REGION Network 83
   RUNG wire#powerrail
      Move(in := "Carrier_54_G120DControlWord", out1 => "DB402_SDC_CARRIER_DRIVE_DATA".Drive_Data.CARRIER[54].Drive_Control)
      Move(in := "Carrier_54_G120DStatusWord", out1 => "DB402_SDC_CARRIER_DRIVE_DATA".Drive_Data.CARRIER[54].Drive_Status)
   END_RUNG
   // the same network as SCL:
   "DB402_SDC_CARRIER_DRIVE_DATA".Drive_Data.CARRIER[54].Drive_Control := "Carrier_54_G120DControlWord";
   "DB402_SDC_CARRIER_DRIVE_DATA".Drive_Data.CARRIER[54].Drive_Status := "Carrier_54_G120DStatusWord";
END_REGION

REGION Network 84
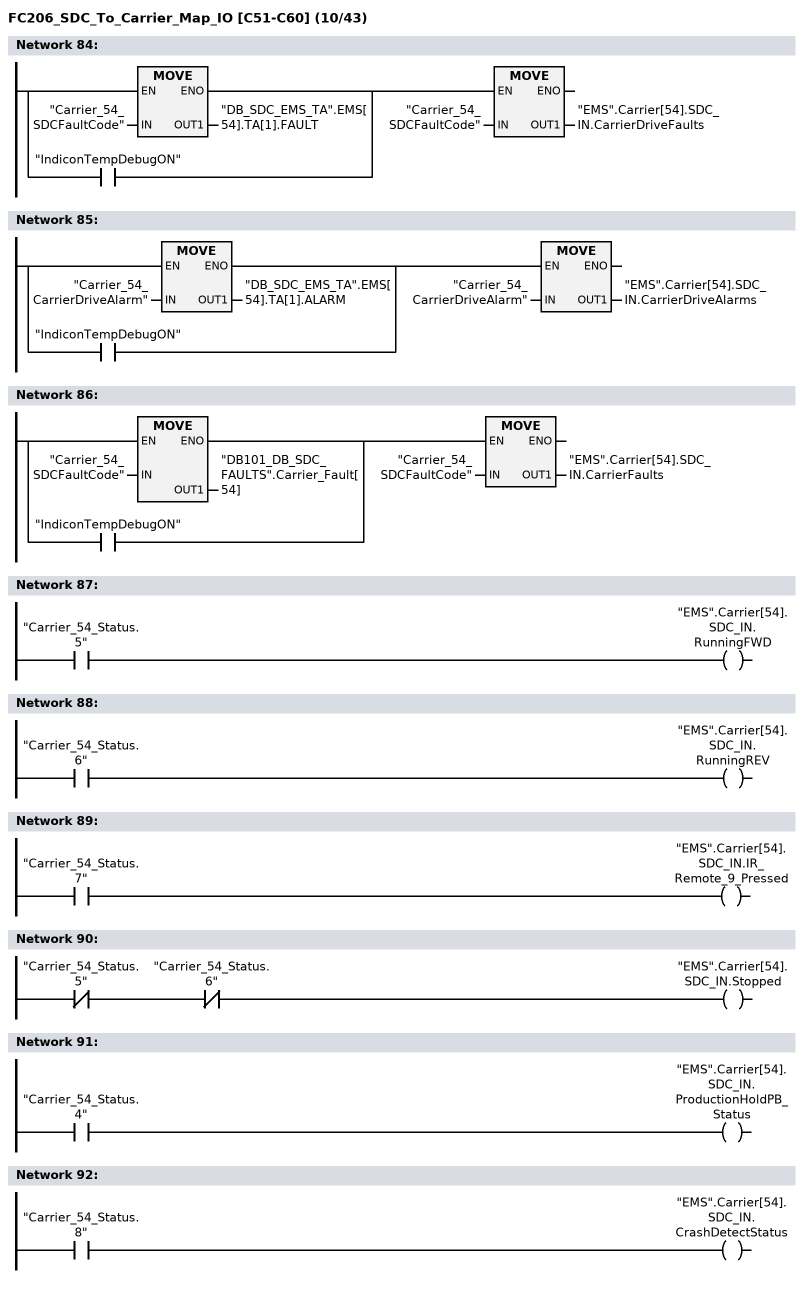
   RUNG wire#powerrail
      Move(in := "Carrier_54_SDCFaultCode", out1 => "DB_SDC_EMS_TA".EMS[54].TA[1].FAULT)
      wire#w1
      Move(in := "Carrier_54_SDCFaultCode", out1 => "EMS".Carrier[54].SDC_IN.CarrierDriveFaults)
   END_RUNG
   RUNG wire#powerrail
      Contact( "IndiconTempDebugON" )
   END_RUNG wire#w1
   // the same network as SCL:
   "DB_SDC_EMS_TA".EMS[54].TA[1].FAULT := "Carrier_54_SDCFaultCode";
   IF TRUE OR "IndiconTempDebugON" THEN
       "EMS".Carrier[54].SDC_IN.CarrierDriveFaults := "Carrier_54_SDCFaultCode";
   END_IF;
END_REGION

REGION Network 85
   RUNG wire#powerrail
      Move(in := "Carrier_54_CarrierDriveAlarm", out1 => "DB_SDC_EMS_TA".EMS[54].TA[1].ALARM)
      wire#w1
      Move(in := "Carrier_54_CarrierDriveAlarm", out1 => "EMS".Carrier[54].SDC_IN.CarrierDriveAlarms)
   END_RUNG
   RUNG wire#powerrail
      Contact( "IndiconTempDebugON" )
   END_RUNG wire#w1
   // the same network as SCL:
   "DB_SDC_EMS_TA".EMS[54].TA[1].ALARM := "Carrier_54_CarrierDriveAlarm";
   IF TRUE OR "IndiconTempDebugON" THEN
       "EMS".Carrier[54].SDC_IN.CarrierDriveAlarms := "Carrier_54_CarrierDriveAlarm";
   END_IF;
END_REGION

REGION Network 86
   RUNG wire#powerrail
      Move(in := "Carrier_54_SDCFaultCode", out1 => "DB101_DB_SDC_FAULTS".Carrier_Fault[54])
      wire#w1
      Move(in := "Carrier_54_SDCFaultCode", out1 => "EMS".Carrier[54].SDC_IN.CarrierFaults)
   END_RUNG
   RUNG wire#powerrail
      Contact( "IndiconTempDebugON" )
   END_RUNG wire#w1
   // the same network as SCL:
   "DB101_DB_SDC_FAULTS".Carrier_Fault[54] := "Carrier_54_SDCFaultCode";
   IF TRUE OR "IndiconTempDebugON" THEN
       "EMS".Carrier[54].SDC_IN.CarrierFaults := "Carrier_54_SDCFaultCode";
   END_IF;
END_REGION

REGION Network 87
   RUNG wire#powerrail
      Contact( "Carrier_54_Status.5" )
      Coil( "EMS".Carrier[54].SDC_IN.RunningFWD )
   END_RUNG
   // the same network as SCL:
   "EMS".Carrier[54].SDC_IN.RunningFWD := "Carrier_54_Status.5";
END_REGION

REGION Network 88
   RUNG wire#powerrail
      Contact( "Carrier_54_Status.6" )
      Coil( "EMS".Carrier[54].SDC_IN.RunningREV )
   END_RUNG
   // the same network as SCL:
   "EMS".Carrier[54].SDC_IN.RunningREV := "Carrier_54_Status.6";
END_REGION

REGION Network 89
   RUNG wire#powerrail
      Contact( "Carrier_54_Status.7" )
      Coil( "EMS".Carrier[54].SDC_IN.IR_Remote_9_Pressed )
   END_RUNG
   // the same network as SCL:
   "EMS".Carrier[54].SDC_IN.IR_Remote_9_Pressed := "Carrier_54_Status.7";
END_REGION

REGION Network 90
   RUNG wire#powerrail
      I_Contact( "Carrier_54_Status.5" )
      I_Contact( "Carrier_54_Status.6" )
      Coil( "EMS".Carrier[54].SDC_IN.Stopped )
   END_RUNG
   // the same network as SCL:
   "EMS".Carrier[54].SDC_IN.Stopped := NOT "Carrier_54_Status.5" AND NOT "Carrier_54_Status.6";
END_REGION

REGION Network 91
   RUNG wire#powerrail
      Contact( "Carrier_54_Status.4" )
      Coil( "EMS".Carrier[54].SDC_IN.ProductionHoldPB_Status )
   END_RUNG
   // the same network as SCL:
   "EMS".Carrier[54].SDC_IN.ProductionHoldPB_Status := "Carrier_54_Status.4";
END_REGION

REGION Network 92
   RUNG wire#powerrail
      Contact( "Carrier_54_Status.8" )
      Coil( "EMS".Carrier[54].SDC_IN.CrashDetectStatus )
   END_RUNG
   // the same network as SCL:
   "EMS".Carrier[54].SDC_IN.CrashDetectStatus := "Carrier_54_Status.8";
END_REGION

REGION Network 93
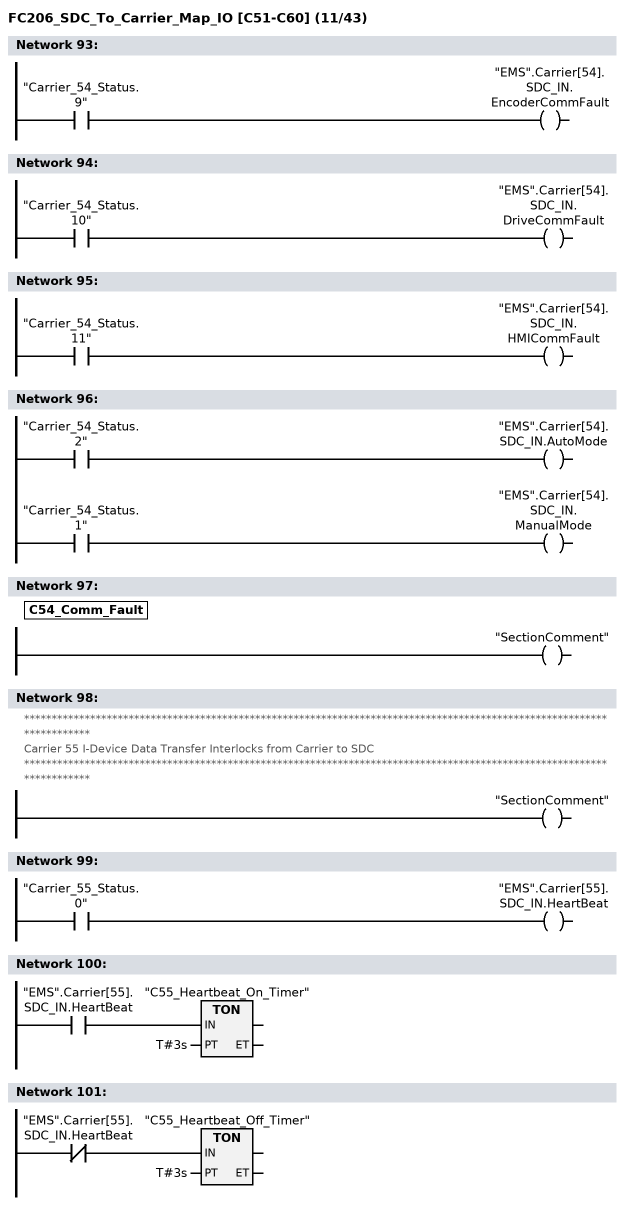
   RUNG wire#powerrail
      Contact( "Carrier_54_Status.9" )
      Coil( "EMS".Carrier[54].SDC_IN.EncoderCommFault )
   END_RUNG
   // the same network as SCL:
   "EMS".Carrier[54].SDC_IN.EncoderCommFault := "Carrier_54_Status.9";
END_REGION

REGION Network 94
   RUNG wire#powerrail
      Contact( "Carrier_54_Status.10" )
      Coil( "EMS".Carrier[54].SDC_IN.DriveCommFault )
   END_RUNG
   // the same network as SCL:
   "EMS".Carrier[54].SDC_IN.DriveCommFault := "Carrier_54_Status.10";
END_REGION

REGION Network 95
   RUNG wire#powerrail
      Contact( "Carrier_54_Status.11" )
      Coil( "EMS".Carrier[54].SDC_IN.HMICommFault )
   END_RUNG
   // the same network as SCL:
   "EMS".Carrier[54].SDC_IN.HMICommFault := "Carrier_54_Status.11";
END_REGION

REGION Network 96
   RUNG wire#powerrail
      Contact( "Carrier_54_Status.2" )
      Coil( "EMS".Carrier[54].SDC_IN.AutoMode )
   END_RUNG
   RUNG wire#powerrail
      Contact( "Carrier_54_Status.1" )
      Coil( "EMS".Carrier[54].SDC_IN.ManualMode )
   END_RUNG
   // the same network as SCL:
   "EMS".Carrier[54].SDC_IN.AutoMode := "Carrier_54_Status.2";
   "EMS".Carrier[54].SDC_IN.ManualMode := "Carrier_54_Status.1";
END_REGION

REGION Network 97
   Label( C54_Comm_Fault )
   RUNG wire#powerrail
      Coil( "SectionComment" )
   END_RUNG
   // the same network as SCL:
   C54_Comm_Fault:
   "SectionComment" := TRUE;
END_REGION

REGION Network 98
   // **********************************************************************************************************************
   // 
   // Carrier 55 I-Device Data Transfer Interlocks from Carrier to SDC
   // 
   // **********************************************************************************************************************
   RUNG wire#powerrail
      Coil( "SectionComment" )
   END_RUNG
   // the same network as SCL:
   "SectionComment" := TRUE;
END_REGION

REGION Network 99
   RUNG wire#powerrail
      Contact( "Carrier_55_Status.0" )
      Coil( "EMS".Carrier[55].SDC_IN.HeartBeat )
   END_RUNG
   // the same network as SCL:
   "EMS".Carrier[55].SDC_IN.HeartBeat := "Carrier_55_Status.0";
END_REGION

REGION Network 100
   "C55_Heartbeat_On_Timer".TON(IN := "EMS".Carrier[55].SDC_IN.HeartBeat, PT := T#3s);
END_REGION

REGION Network 101
   "C55_Heartbeat_Off_Timer".TON(IN := NOT "EMS".Carrier[55].SDC_IN.HeartBeat, PT := T#3s);
END_REGION

REGION Network 102
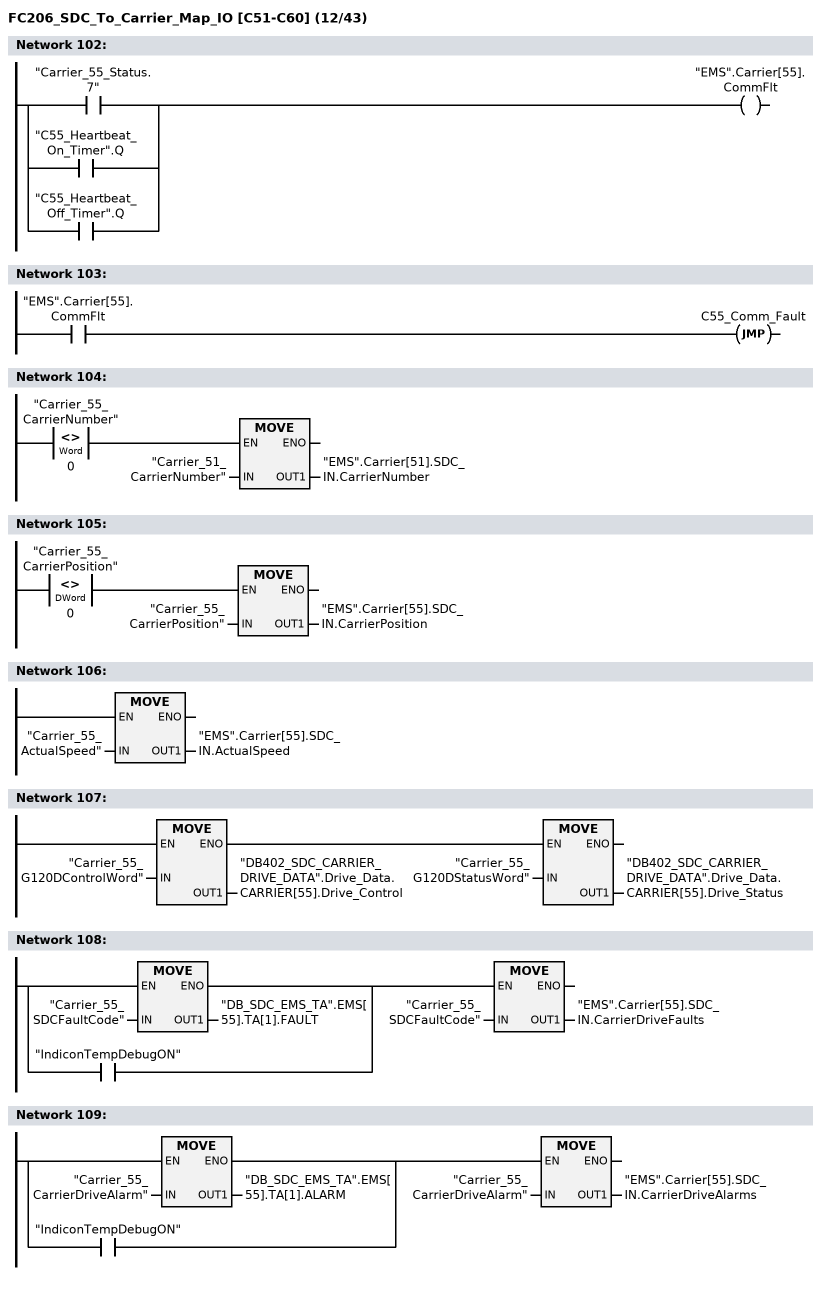
   RUNG wire#powerrail
      Contact( "Carrier_55_Status.7" )
      wire#w1
      Coil( "EMS".Carrier[55].CommFlt )
   END_RUNG
   RUNG wire#powerrail
      Contact( "C55_Heartbeat_On_Timer".Q )
   END_RUNG wire#w1
   RUNG wire#powerrail
      Contact( "C55_Heartbeat_Off_Timer".Q )
   END_RUNG wire#w1
   // the same network as SCL:
   "EMS".Carrier[55].CommFlt := "Carrier_55_Status.7" OR "C55_Heartbeat_On_Timer".Q OR "C55_Heartbeat_Off_Timer".Q;
END_REGION

REGION Network 103
   RUNG wire#powerrail
      Contact( "EMS".Carrier[55].CommFlt )
      JumpCoil( C55_Comm_Fault )
   END_RUNG
   // the same network as SCL:
   IF "EMS".Carrier[55].CommFlt THEN GOTO C55_Comm_Fault; END_IF;
END_REGION

REGION Network 104
   RUNG wire#powerrail
      { S7_Templates := "SrcType := Word" } NE_Contact(in1 := "Carrier_55_CarrierNumber", in2 := 0)
      Move(in := "Carrier_51_CarrierNumber", out1 => "EMS".Carrier[51].SDC_IN.CarrierNumber)
   END_RUNG
   // the same network as SCL:
   IF "Carrier_55_CarrierNumber" <> 0 THEN
       "EMS".Carrier[51].SDC_IN.CarrierNumber := "Carrier_51_CarrierNumber";
   END_IF;
END_REGION

REGION Network 105
   RUNG wire#powerrail
      { S7_Templates := "SrcType := DWord" } NE_Contact(in1 := "Carrier_55_CarrierPosition", in2 := 0)
      Move(in := "Carrier_55_CarrierPosition", out1 => "EMS".Carrier[55].SDC_IN.CarrierPosition)
   END_RUNG
   // the same network as SCL:
   IF "Carrier_55_CarrierPosition" <> 0 THEN
       "EMS".Carrier[55].SDC_IN.CarrierPosition := "Carrier_55_CarrierPosition";
   END_IF;
END_REGION

REGION Network 106
   RUNG wire#powerrail
      Move(in := "Carrier_55_ActualSpeed", out1 => "EMS".Carrier[55].SDC_IN.ActualSpeed)
   END_RUNG
   // the same network as SCL:
   "EMS".Carrier[55].SDC_IN.ActualSpeed := "Carrier_55_ActualSpeed";
END_REGION

REGION Network 107
   RUNG wire#powerrail
      Move(in := "Carrier_55_G120DControlWord", out1 => "DB402_SDC_CARRIER_DRIVE_DATA".Drive_Data.CARRIER[55].Drive_Control)
      Move(in := "Carrier_55_G120DStatusWord", out1 => "DB402_SDC_CARRIER_DRIVE_DATA".Drive_Data.CARRIER[55].Drive_Status)
   END_RUNG
   // the same network as SCL:
   "DB402_SDC_CARRIER_DRIVE_DATA".Drive_Data.CARRIER[55].Drive_Control := "Carrier_55_G120DControlWord";
   "DB402_SDC_CARRIER_DRIVE_DATA".Drive_Data.CARRIER[55].Drive_Status := "Carrier_55_G120DStatusWord";
END_REGION

REGION Network 108
   RUNG wire#powerrail
      Move(in := "Carrier_55_SDCFaultCode", out1 => "DB_SDC_EMS_TA".EMS[55].TA[1].FAULT)
      wire#w1
      Move(in := "Carrier_55_SDCFaultCode", out1 => "EMS".Carrier[55].SDC_IN.CarrierDriveFaults)
   END_RUNG
   RUNG wire#powerrail
      Contact( "IndiconTempDebugON" )
   END_RUNG wire#w1
   // the same network as SCL:
   "DB_SDC_EMS_TA".EMS[55].TA[1].FAULT := "Carrier_55_SDCFaultCode";
   IF TRUE OR "IndiconTempDebugON" THEN
       "EMS".Carrier[55].SDC_IN.CarrierDriveFaults := "Carrier_55_SDCFaultCode";
   END_IF;
END_REGION

REGION Network 109
   RUNG wire#powerrail
      Move(in := "Carrier_55_CarrierDriveAlarm", out1 => "DB_SDC_EMS_TA".EMS[55].TA[1].ALARM)
      wire#w1
      Move(in := "Carrier_55_CarrierDriveAlarm", out1 => "EMS".Carrier[55].SDC_IN.CarrierDriveAlarms)
   END_RUNG
   RUNG wire#powerrail
      Contact( "IndiconTempDebugON" )
   END_RUNG wire#w1
   // the same network as SCL:
   "DB_SDC_EMS_TA".EMS[55].TA[1].ALARM := "Carrier_55_CarrierDriveAlarm";
   IF TRUE OR "IndiconTempDebugON" THEN
       "EMS".Carrier[55].SDC_IN.CarrierDriveAlarms := "Carrier_55_CarrierDriveAlarm";
   END_IF;
END_REGION

REGION Network 110
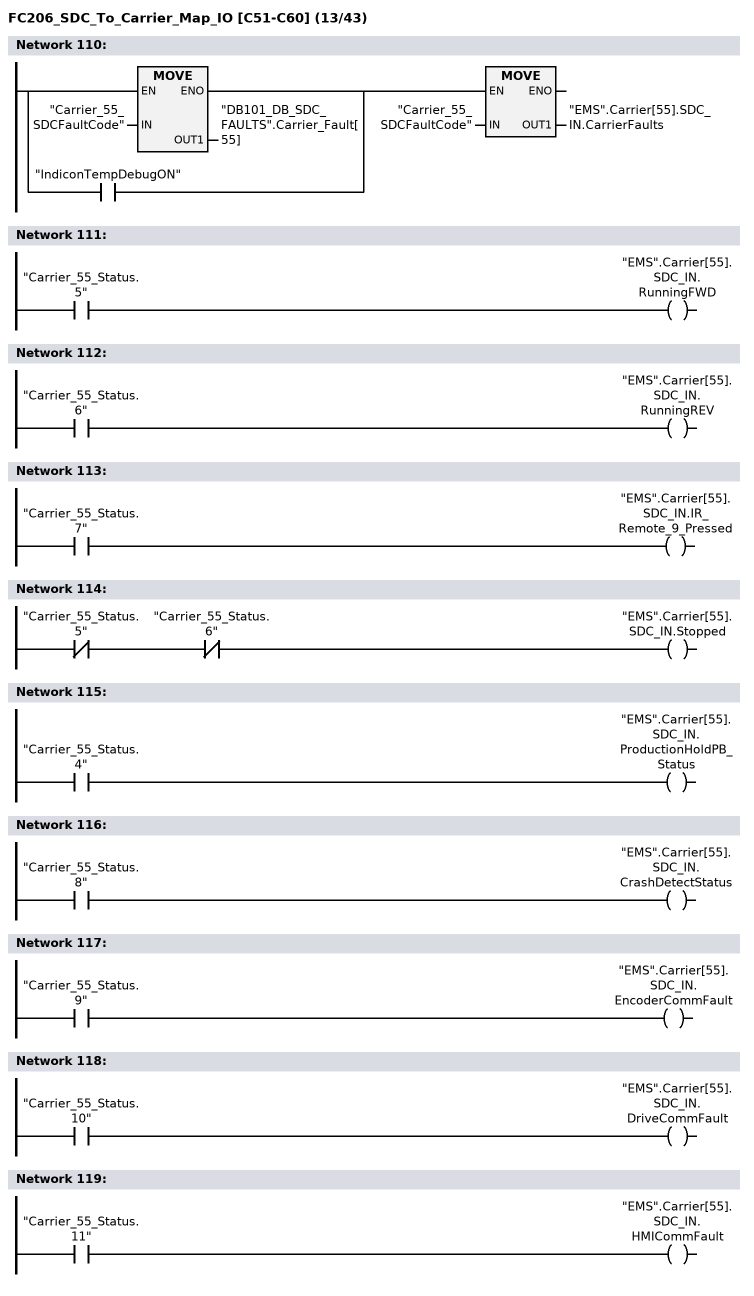
   RUNG wire#powerrail
      Move(in := "Carrier_55_SDCFaultCode", out1 => "DB101_DB_SDC_FAULTS".Carrier_Fault[55])
      wire#w1
      Move(in := "Carrier_55_SDCFaultCode", out1 => "EMS".Carrier[55].SDC_IN.CarrierFaults)
   END_RUNG
   RUNG wire#powerrail
      Contact( "IndiconTempDebugON" )
   END_RUNG wire#w1
   // the same network as SCL:
   "DB101_DB_SDC_FAULTS".Carrier_Fault[55] := "Carrier_55_SDCFaultCode";
   IF TRUE OR "IndiconTempDebugON" THEN
       "EMS".Carrier[55].SDC_IN.CarrierFaults := "Carrier_55_SDCFaultCode";
   END_IF;
END_REGION

REGION Network 111
   RUNG wire#powerrail
      Contact( "Carrier_55_Status.5" )
      Coil( "EMS".Carrier[55].SDC_IN.RunningFWD )
   END_RUNG
   // the same network as SCL:
   "EMS".Carrier[55].SDC_IN.RunningFWD := "Carrier_55_Status.5";
END_REGION

REGION Network 112
   RUNG wire#powerrail
      Contact( "Carrier_55_Status.6" )
      Coil( "EMS".Carrier[55].SDC_IN.RunningREV )
   END_RUNG
   // the same network as SCL:
   "EMS".Carrier[55].SDC_IN.RunningREV := "Carrier_55_Status.6";
END_REGION

REGION Network 113
   RUNG wire#powerrail
      Contact( "Carrier_55_Status.7" )
      Coil( "EMS".Carrier[55].SDC_IN.IR_Remote_9_Pressed )
   END_RUNG
   // the same network as SCL:
   "EMS".Carrier[55].SDC_IN.IR_Remote_9_Pressed := "Carrier_55_Status.7";
END_REGION

REGION Network 114
   RUNG wire#powerrail
      I_Contact( "Carrier_55_Status.5" )
      I_Contact( "Carrier_55_Status.6" )
      Coil( "EMS".Carrier[55].SDC_IN.Stopped )
   END_RUNG
   // the same network as SCL:
   "EMS".Carrier[55].SDC_IN.Stopped := NOT "Carrier_55_Status.5" AND NOT "Carrier_55_Status.6";
END_REGION

REGION Network 115
   RUNG wire#powerrail
      Contact( "Carrier_55_Status.4" )
      Coil( "EMS".Carrier[55].SDC_IN.ProductionHoldPB_Status )
   END_RUNG
   // the same network as SCL:
   "EMS".Carrier[55].SDC_IN.ProductionHoldPB_Status := "Carrier_55_Status.4";
END_REGION

REGION Network 116
   RUNG wire#powerrail
      Contact( "Carrier_55_Status.8" )
      Coil( "EMS".Carrier[55].SDC_IN.CrashDetectStatus )
   END_RUNG
   // the same network as SCL:
   "EMS".Carrier[55].SDC_IN.CrashDetectStatus := "Carrier_55_Status.8";
END_REGION

REGION Network 117
   RUNG wire#powerrail
      Contact( "Carrier_55_Status.9" )
      Coil( "EMS".Carrier[55].SDC_IN.EncoderCommFault )
   END_RUNG
   // the same network as SCL:
   "EMS".Carrier[55].SDC_IN.EncoderCommFault := "Carrier_55_Status.9";
END_REGION

REGION Network 118
   RUNG wire#powerrail
      Contact( "Carrier_55_Status.10" )
      Coil( "EMS".Carrier[55].SDC_IN.DriveCommFault )
   END_RUNG
   // the same network as SCL:
   "EMS".Carrier[55].SDC_IN.DriveCommFault := "Carrier_55_Status.10";
END_REGION

REGION Network 119
   RUNG wire#powerrail
      Contact( "Carrier_55_Status.11" )
      Coil( "EMS".Carrier[55].SDC_IN.HMICommFault )
   END_RUNG
   // the same network as SCL:
   "EMS".Carrier[55].SDC_IN.HMICommFault := "Carrier_55_Status.11";
END_REGION

REGION Network 120
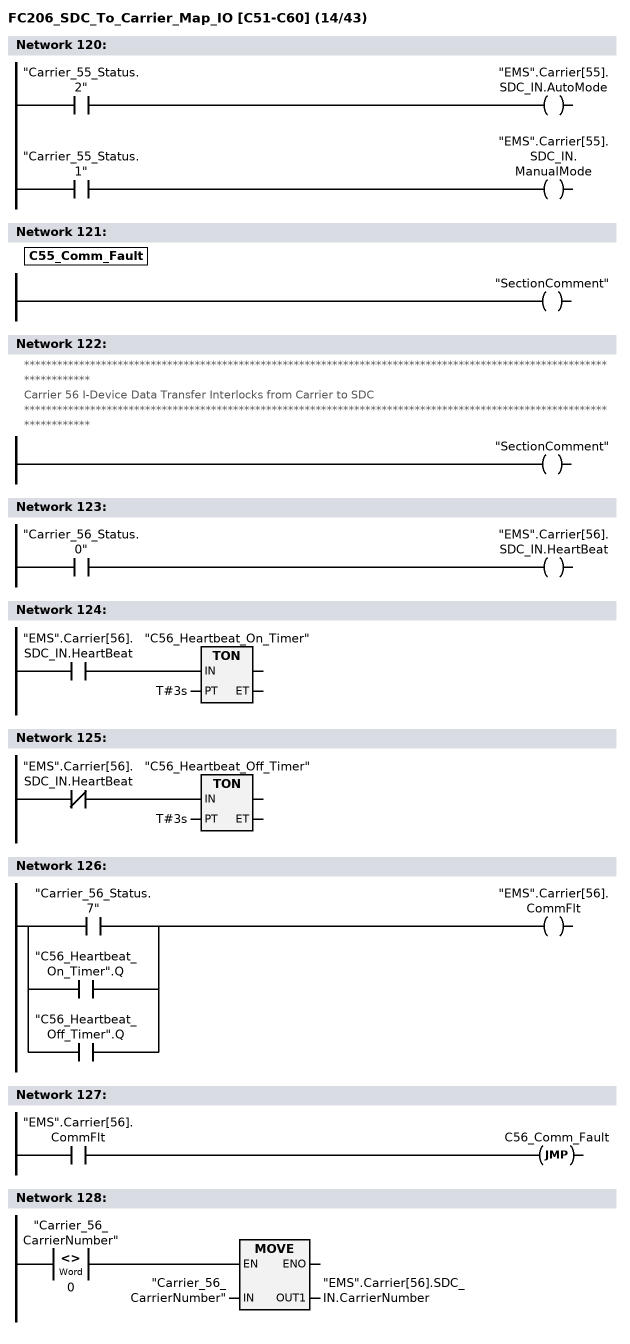
   RUNG wire#powerrail
      Contact( "Carrier_55_Status.2" )
      Coil( "EMS".Carrier[55].SDC_IN.AutoMode )
   END_RUNG
   RUNG wire#powerrail
      Contact( "Carrier_55_Status.1" )
      Coil( "EMS".Carrier[55].SDC_IN.ManualMode )
   END_RUNG
   // the same network as SCL:
   "EMS".Carrier[55].SDC_IN.AutoMode := "Carrier_55_Status.2";
   "EMS".Carrier[55].SDC_IN.ManualMode := "Carrier_55_Status.1";
END_REGION

REGION Network 121
   Label( C55_Comm_Fault )
   RUNG wire#powerrail
      Coil( "SectionComment" )
   END_RUNG
   // the same network as SCL:
   C55_Comm_Fault:
   "SectionComment" := TRUE;
END_REGION

REGION Network 122
   // **********************************************************************************************************************
   // 
   // Carrier 56 I-Device Data Transfer Interlocks from Carrier to SDC
   // 
   // **********************************************************************************************************************
   RUNG wire#powerrail
      Coil( "SectionComment" )
   END_RUNG
   // the same network as SCL:
   "SectionComment" := TRUE;
END_REGION

REGION Network 123
   RUNG wire#powerrail
      Contact( "Carrier_56_Status.0" )
      Coil( "EMS".Carrier[56].SDC_IN.HeartBeat )
   END_RUNG
   // the same network as SCL:
   "EMS".Carrier[56].SDC_IN.HeartBeat := "Carrier_56_Status.0";
END_REGION

REGION Network 124
   "C56_Heartbeat_On_Timer".TON(IN := "EMS".Carrier[56].SDC_IN.HeartBeat, PT := T#3s);
END_REGION

REGION Network 125
   "C56_Heartbeat_Off_Timer".TON(IN := NOT "EMS".Carrier[56].SDC_IN.HeartBeat, PT := T#3s);
END_REGION

REGION Network 126
   RUNG wire#powerrail
      Contact( "Carrier_56_Status.7" )
      wire#w1
      Coil( "EMS".Carrier[56].CommFlt )
   END_RUNG
   RUNG wire#powerrail
      Contact( "C56_Heartbeat_On_Timer".Q )
   END_RUNG wire#w1
   RUNG wire#powerrail
      Contact( "C56_Heartbeat_Off_Timer".Q )
   END_RUNG wire#w1
   // the same network as SCL:
   "EMS".Carrier[56].CommFlt := "Carrier_56_Status.7" OR "C56_Heartbeat_On_Timer".Q OR "C56_Heartbeat_Off_Timer".Q;
END_REGION

REGION Network 127
   RUNG wire#powerrail
      Contact( "EMS".Carrier[56].CommFlt )
      JumpCoil( C56_Comm_Fault )
   END_RUNG
   // the same network as SCL:
   IF "EMS".Carrier[56].CommFlt THEN GOTO C56_Comm_Fault; END_IF;
END_REGION

REGION Network 128
   RUNG wire#powerrail
      { S7_Templates := "SrcType := Word" } NE_Contact(in1 := "Carrier_56_CarrierNumber", in2 := 0)
      Move(in := "Carrier_56_CarrierNumber", out1 => "EMS".Carrier[56].SDC_IN.CarrierNumber)
   END_RUNG
   // the same network as SCL:
   IF "Carrier_56_CarrierNumber" <> 0 THEN
       "EMS".Carrier[56].SDC_IN.CarrierNumber := "Carrier_56_CarrierNumber";
   END_IF;
END_REGION

REGION Network 129
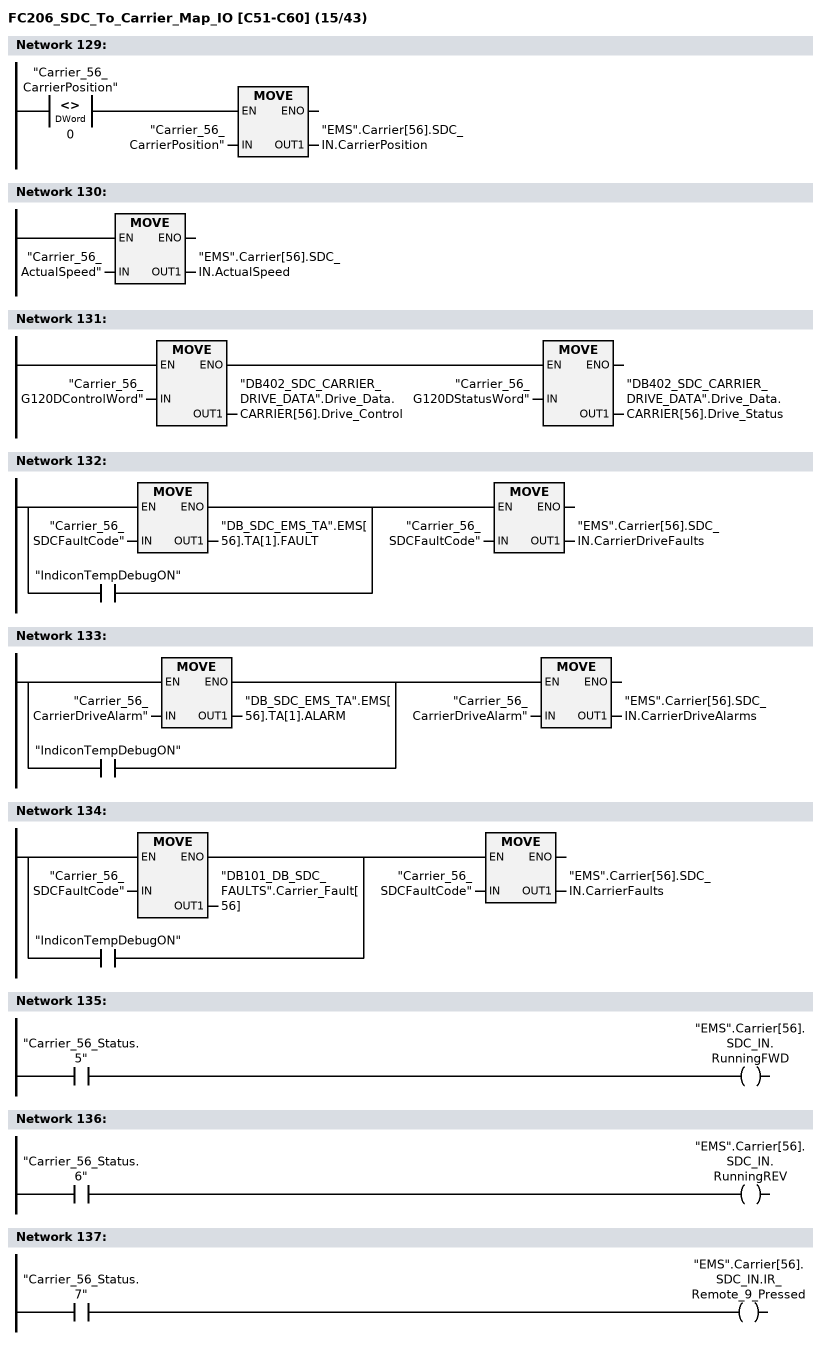
   RUNG wire#powerrail
      { S7_Templates := "SrcType := DWord" } NE_Contact(in1 := "Carrier_56_CarrierPosition", in2 := 0)
      Move(in := "Carrier_56_CarrierPosition", out1 => "EMS".Carrier[56].SDC_IN.CarrierPosition)
   END_RUNG
   // the same network as SCL:
   IF "Carrier_56_CarrierPosition" <> 0 THEN
       "EMS".Carrier[56].SDC_IN.CarrierPosition := "Carrier_56_CarrierPosition";
   END_IF;
END_REGION

REGION Network 130
   RUNG wire#powerrail
      Move(in := "Carrier_56_ActualSpeed", out1 => "EMS".Carrier[56].SDC_IN.ActualSpeed)
   END_RUNG
   // the same network as SCL:
   "EMS".Carrier[56].SDC_IN.ActualSpeed := "Carrier_56_ActualSpeed";
END_REGION

REGION Network 131
   RUNG wire#powerrail
      Move(in := "Carrier_56_G120DControlWord", out1 => "DB402_SDC_CARRIER_DRIVE_DATA".Drive_Data.CARRIER[56].Drive_Control)
      Move(in := "Carrier_56_G120DStatusWord", out1 => "DB402_SDC_CARRIER_DRIVE_DATA".Drive_Data.CARRIER[56].Drive_Status)
   END_RUNG
   // the same network as SCL:
   "DB402_SDC_CARRIER_DRIVE_DATA".Drive_Data.CARRIER[56].Drive_Control := "Carrier_56_G120DControlWord";
   "DB402_SDC_CARRIER_DRIVE_DATA".Drive_Data.CARRIER[56].Drive_Status := "Carrier_56_G120DStatusWord";
END_REGION

REGION Network 132
   RUNG wire#powerrail
      Move(in := "Carrier_56_SDCFaultCode", out1 => "DB_SDC_EMS_TA".EMS[56].TA[1].FAULT)
      wire#w1
      Move(in := "Carrier_56_SDCFaultCode", out1 => "EMS".Carrier[56].SDC_IN.CarrierDriveFaults)
   END_RUNG
   RUNG wire#powerrail
      Contact( "IndiconTempDebugON" )
   END_RUNG wire#w1
   // the same network as SCL:
   "DB_SDC_EMS_TA".EMS[56].TA[1].FAULT := "Carrier_56_SDCFaultCode";
   IF TRUE OR "IndiconTempDebugON" THEN
       "EMS".Carrier[56].SDC_IN.CarrierDriveFaults := "Carrier_56_SDCFaultCode";
   END_IF;
END_REGION

REGION Network 133
   RUNG wire#powerrail
      Move(in := "Carrier_56_CarrierDriveAlarm", out1 => "DB_SDC_EMS_TA".EMS[56].TA[1].ALARM)
      wire#w1
      Move(in := "Carrier_56_CarrierDriveAlarm", out1 => "EMS".Carrier[56].SDC_IN.CarrierDriveAlarms)
   END_RUNG
   RUNG wire#powerrail
      Contact( "IndiconTempDebugON" )
   END_RUNG wire#w1
   // the same network as SCL:
   "DB_SDC_EMS_TA".EMS[56].TA[1].ALARM := "Carrier_56_CarrierDriveAlarm";
   IF TRUE OR "IndiconTempDebugON" THEN
       "EMS".Carrier[56].SDC_IN.CarrierDriveAlarms := "Carrier_56_CarrierDriveAlarm";
   END_IF;
END_REGION

REGION Network 134
   RUNG wire#powerrail
      Move(in := "Carrier_56_SDCFaultCode", out1 => "DB101_DB_SDC_FAULTS".Carrier_Fault[56])
      wire#w1
      Move(in := "Carrier_56_SDCFaultCode", out1 => "EMS".Carrier[56].SDC_IN.CarrierFaults)
   END_RUNG
   RUNG wire#powerrail
      Contact( "IndiconTempDebugON" )
   END_RUNG wire#w1
   // the same network as SCL:
   "DB101_DB_SDC_FAULTS".Carrier_Fault[56] := "Carrier_56_SDCFaultCode";
   IF TRUE OR "IndiconTempDebugON" THEN
       "EMS".Carrier[56].SDC_IN.CarrierFaults := "Carrier_56_SDCFaultCode";
   END_IF;
END_REGION

REGION Network 135
   RUNG wire#powerrail
      Contact( "Carrier_56_Status.5" )
      Coil( "EMS".Carrier[56].SDC_IN.RunningFWD )
   END_RUNG
   // the same network as SCL:
   "EMS".Carrier[56].SDC_IN.RunningFWD := "Carrier_56_Status.5";
END_REGION

REGION Network 136
   RUNG wire#powerrail
      Contact( "Carrier_56_Status.6" )
      Coil( "EMS".Carrier[56].SDC_IN.RunningREV )
   END_RUNG
   // the same network as SCL:
   "EMS".Carrier[56].SDC_IN.RunningREV := "Carrier_56_Status.6";
END_REGION

REGION Network 137
   RUNG wire#powerrail
      Contact( "Carrier_56_Status.7" )
      Coil( "EMS".Carrier[56].SDC_IN.IR_Remote_9_Pressed )
   END_RUNG
   // the same network as SCL:
   "EMS".Carrier[56].SDC_IN.IR_Remote_9_Pressed := "Carrier_56_Status.7";
END_REGION

REGION Network 138
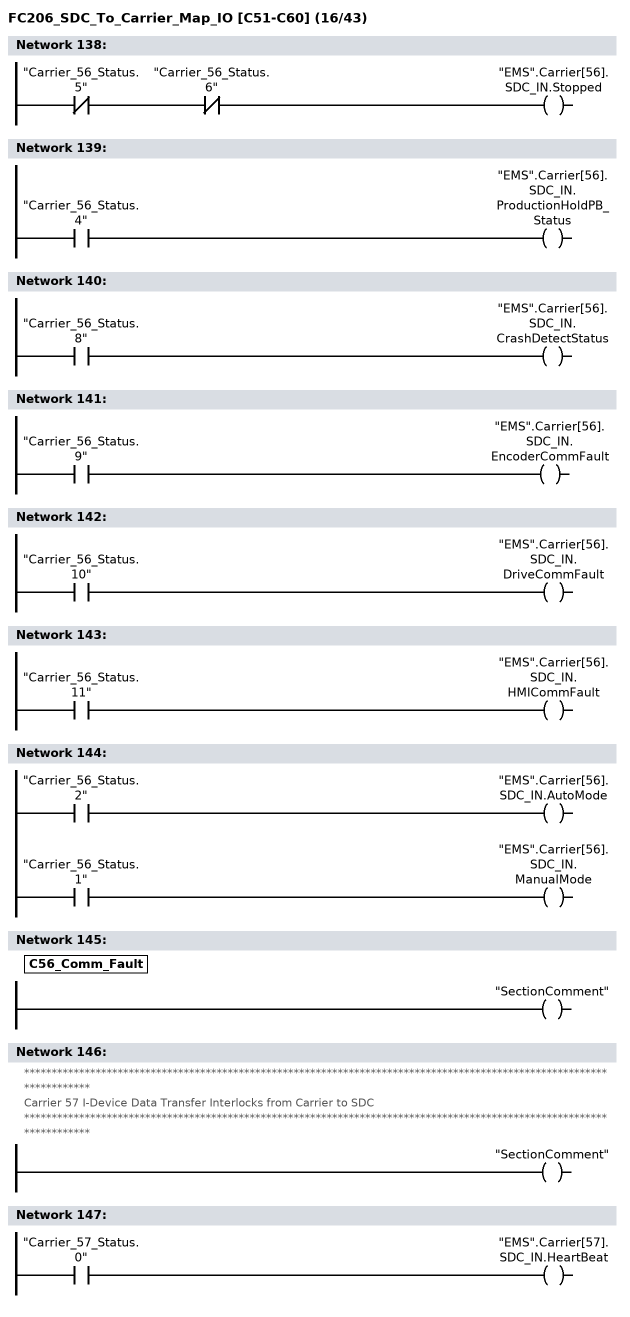
   RUNG wire#powerrail
      I_Contact( "Carrier_56_Status.5" )
      I_Contact( "Carrier_56_Status.6" )
      Coil( "EMS".Carrier[56].SDC_IN.Stopped )
   END_RUNG
   // the same network as SCL:
   "EMS".Carrier[56].SDC_IN.Stopped := NOT "Carrier_56_Status.5" AND NOT "Carrier_56_Status.6";
END_REGION

REGION Network 139
   RUNG wire#powerrail
      Contact( "Carrier_56_Status.4" )
      Coil( "EMS".Carrier[56].SDC_IN.ProductionHoldPB_Status )
   END_RUNG
   // the same network as SCL:
   "EMS".Carrier[56].SDC_IN.ProductionHoldPB_Status := "Carrier_56_Status.4";
END_REGION

REGION Network 140
   RUNG wire#powerrail
      Contact( "Carrier_56_Status.8" )
      Coil( "EMS".Carrier[56].SDC_IN.CrashDetectStatus )
   END_RUNG
   // the same network as SCL:
   "EMS".Carrier[56].SDC_IN.CrashDetectStatus := "Carrier_56_Status.8";
END_REGION

REGION Network 141
   RUNG wire#powerrail
      Contact( "Carrier_56_Status.9" )
      Coil( "EMS".Carrier[56].SDC_IN.EncoderCommFault )
   END_RUNG
   // the same network as SCL:
   "EMS".Carrier[56].SDC_IN.EncoderCommFault := "Carrier_56_Status.9";
END_REGION

REGION Network 142
   RUNG wire#powerrail
      Contact( "Carrier_56_Status.10" )
      Coil( "EMS".Carrier[56].SDC_IN.DriveCommFault )
   END_RUNG
   // the same network as SCL:
   "EMS".Carrier[56].SDC_IN.DriveCommFault := "Carrier_56_Status.10";
END_REGION

REGION Network 143
   RUNG wire#powerrail
      Contact( "Carrier_56_Status.11" )
      Coil( "EMS".Carrier[56].SDC_IN.HMICommFault )
   END_RUNG
   // the same network as SCL:
   "EMS".Carrier[56].SDC_IN.HMICommFault := "Carrier_56_Status.11";
END_REGION

REGION Network 144
   RUNG wire#powerrail
      Contact( "Carrier_56_Status.2" )
      Coil( "EMS".Carrier[56].SDC_IN.AutoMode )
   END_RUNG
   RUNG wire#powerrail
      Contact( "Carrier_56_Status.1" )
      Coil( "EMS".Carrier[56].SDC_IN.ManualMode )
   END_RUNG
   // the same network as SCL:
   "EMS".Carrier[56].SDC_IN.AutoMode := "Carrier_56_Status.2";
   "EMS".Carrier[56].SDC_IN.ManualMode := "Carrier_56_Status.1";
END_REGION

REGION Network 145
   Label( C56_Comm_Fault )
   RUNG wire#powerrail
      Coil( "SectionComment" )
   END_RUNG
   // the same network as SCL:
   C56_Comm_Fault:
   "SectionComment" := TRUE;
END_REGION

REGION Network 146
   // **********************************************************************************************************************
   // 
   // Carrier 57 I-Device Data Transfer Interlocks from Carrier to SDC
   // 
   // **********************************************************************************************************************
   RUNG wire#powerrail
      Coil( "SectionComment" )
   END_RUNG
   // the same network as SCL:
   "SectionComment" := TRUE;
END_REGION

REGION Network 147
   RUNG wire#powerrail
      Contact( "Carrier_57_Status.0" )
      Coil( "EMS".Carrier[57].SDC_IN.HeartBeat )
   END_RUNG
   // the same network as SCL:
   "EMS".Carrier[57].SDC_IN.HeartBeat := "Carrier_57_Status.0";
END_REGION

REGION Network 148
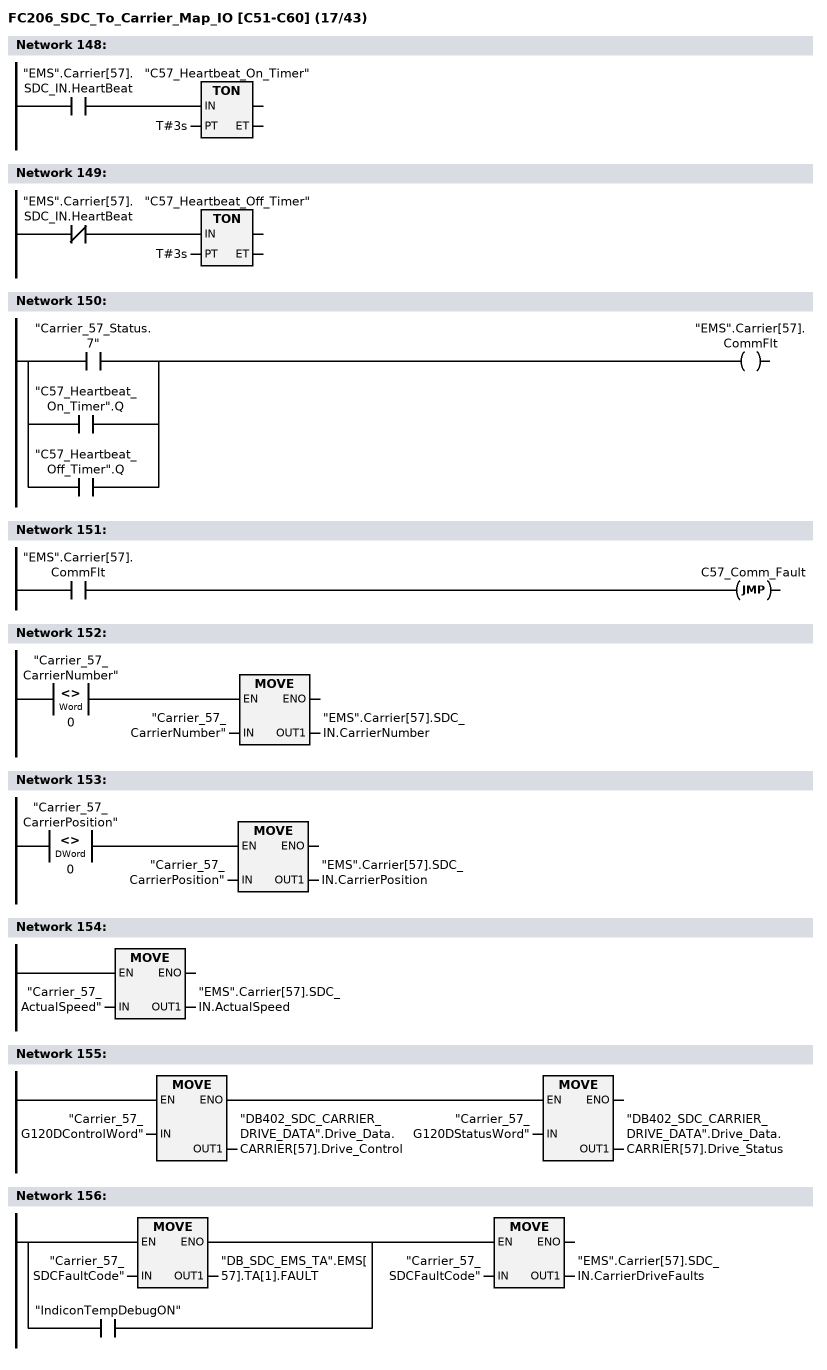
   "C57_Heartbeat_On_Timer".TON(IN := "EMS".Carrier[57].SDC_IN.HeartBeat, PT := T#3s);
END_REGION

REGION Network 149
   "C57_Heartbeat_Off_Timer".TON(IN := NOT "EMS".Carrier[57].SDC_IN.HeartBeat, PT := T#3s);
END_REGION

REGION Network 150
   RUNG wire#powerrail
      Contact( "Carrier_57_Status.7" )
      wire#w1
      Coil( "EMS".Carrier[57].CommFlt )
   END_RUNG
   RUNG wire#powerrail
      Contact( "C57_Heartbeat_On_Timer".Q )
   END_RUNG wire#w1
   RUNG wire#powerrail
      Contact( "C57_Heartbeat_Off_Timer".Q )
   END_RUNG wire#w1
   // the same network as SCL:
   "EMS".Carrier[57].CommFlt := "Carrier_57_Status.7" OR "C57_Heartbeat_On_Timer".Q OR "C57_Heartbeat_Off_Timer".Q;
END_REGION

REGION Network 151
   RUNG wire#powerrail
      Contact( "EMS".Carrier[57].CommFlt )
      JumpCoil( C57_Comm_Fault )
   END_RUNG
   // the same network as SCL:
   IF "EMS".Carrier[57].CommFlt THEN GOTO C57_Comm_Fault; END_IF;
END_REGION

REGION Network 152
   RUNG wire#powerrail
      { S7_Templates := "SrcType := Word" } NE_Contact(in1 := "Carrier_57_CarrierNumber", in2 := 0)
      Move(in := "Carrier_57_CarrierNumber", out1 => "EMS".Carrier[57].SDC_IN.CarrierNumber)
   END_RUNG
   // the same network as SCL:
   IF "Carrier_57_CarrierNumber" <> 0 THEN
       "EMS".Carrier[57].SDC_IN.CarrierNumber := "Carrier_57_CarrierNumber";
   END_IF;
END_REGION

REGION Network 153
   RUNG wire#powerrail
      { S7_Templates := "SrcType := DWord" } NE_Contact(in1 := "Carrier_57_CarrierPosition", in2 := 0)
      Move(in := "Carrier_57_CarrierPosition", out1 => "EMS".Carrier[57].SDC_IN.CarrierPosition)
   END_RUNG
   // the same network as SCL:
   IF "Carrier_57_CarrierPosition" <> 0 THEN
       "EMS".Carrier[57].SDC_IN.CarrierPosition := "Carrier_57_CarrierPosition";
   END_IF;
END_REGION

REGION Network 154
   RUNG wire#powerrail
      Move(in := "Carrier_57_ActualSpeed", out1 => "EMS".Carrier[57].SDC_IN.ActualSpeed)
   END_RUNG
   // the same network as SCL:
   "EMS".Carrier[57].SDC_IN.ActualSpeed := "Carrier_57_ActualSpeed";
END_REGION

REGION Network 155
   RUNG wire#powerrail
      Move(in := "Carrier_57_G120DControlWord", out1 => "DB402_SDC_CARRIER_DRIVE_DATA".Drive_Data.CARRIER[57].Drive_Control)
      Move(in := "Carrier_57_G120DStatusWord", out1 => "DB402_SDC_CARRIER_DRIVE_DATA".Drive_Data.CARRIER[57].Drive_Status)
   END_RUNG
   // the same network as SCL:
   "DB402_SDC_CARRIER_DRIVE_DATA".Drive_Data.CARRIER[57].Drive_Control := "Carrier_57_G120DControlWord";
   "DB402_SDC_CARRIER_DRIVE_DATA".Drive_Data.CARRIER[57].Drive_Status := "Carrier_57_G120DStatusWord";
END_REGION
